screen "08 BTCS MAIN" 1280x800, template "Template"
   Rectangle "Rectangle_2" at 150,205 size 480x40
      Appearance <- "2102_TIME_CALCS_DB_DE_OX_TMR_DN"
   TextField "Text field_7" at 155,210 size 200x30; Text 'De-Oxygenate Time :'
   IOField "I/O field_3" at 360,210 size 60x30; FormatPattern 999
      ProcessValue <- "2110_BTCS_CNTRL_DB_DE_OX_HRS"
   TextField "Text field_8" at 420,210 size 60x30; Text 'Hours'
   IOField "I/O field_4" at 485,210 size 60x30; FormatPattern 99
      ProcessValue <- "2110_BTCS_CNTRL_DB_DE_OX_MINS"
   TextField "Text field_9" at 545,210 size 80x30; Text 'Minutes'
   Rectangle "Rectangle_3" at 150,250 size 480x40
      Appearance <- "2102_TIME_CALCS_DB_DWELL_TMR_DN"
   TextField "Text field_10" at 155,255 size 200x30; Text 'Dwell Time :'
   IOField "I/O field_5" at 360,255 size 60x30; FormatPattern 999
      ProcessValue <- "2110_BTCS_CNTRL_DB_DWELL_HRS"
   TextField "Text field_11" at 420,255 size 60x30; Text 'Hours'
   IOField "I/O field_6" at 485,255 size 60x30; FormatPattern 99
      ProcessValue <- "2110_BTCS_CNTRL_DB_DWELL_MINS"
   TextField "Text field_12" at 545,255 size 80x30; Text 'Minutes'
   Rectangle "Rectangle_4" at 150,295 size 480x40
      Appearance <- "2102_TIME_CALCS_DB_RE_OX_TMR_DN"
   TextField "Text field_13" at 155,300 size 200x30; Text 'Re-Oxygenate Time :'
   IOField "I/O field_7" at 360,300 size 60x30; FormatPattern 999
      ProcessValue <- "2110_BTCS_CNTRL_DB_RE_OX_HRS"
   TextField "Text field_14" at 420,300 size 60x30; Text 'Hours'
   IOField "I/O field_8" at 485,300 size 60x30; FormatPattern 99
      ProcessValue <- "2110_BTCS_CNTRL_DB_RE_OX_MINS"
   TextField "Text field_15" at 545,300 size 80x30; Text 'Minutes'
   Rectangle "Rectangle_5" at 150,340 size 480x40
      Appearance <- "2102_TIME_CALCS_DB_POST_DWELL_TMR_DN"
   TextField "Text field_16" at 155,345 size 200x30; Text 'Post-Dwell Time :'
   IOField "I/O field_9" at 360,345 size 60x30; FormatPattern 999
      ProcessValue <- "2110_BTCS_CNTRL_DB_POST_DWELL_HRS"
   TextField "Text field_17" at 420,345 size 60x30; Text 'Hours'
   IOField "I/O field_10" at 485,345 size 60x30; FormatPattern 99
      ProcessValue <- "2110_BTCS_CNTRL_DB_POST_DWELL_MINS"
   TextField "Text field_18" at 545,345 size 80x30; Text 'Minutes'
   Rectangle "Rectangle_6" at 640,205 size 480x40
      Appearance <- "2102_TIME_CALCS_DB_DE_OX_SP_TMR_DN"
   TextField "Text field_19" at 645,210 size 200x30; Text 'At De-Ox Setpoint :'
   IOField "I/O field_11" at 850,210 size 60x30; FormatPattern 999
      ProcessValue <- "2110_BTCS_CNTRL_DB_DE_OX_SP_HRS"
   TextField "Text field_20" at 910,210 size 60x30; Text 'Hours'
   IOField "I/O field_12" at 975,210 size 60x30; FormatPattern 99
      ProcessValue <- "2110_BTCS_CNTRL_DB_DE_OX_SP_MINS"
   TextField "Text field_21" at 1035,210 size 80x30; Text 'Minutes'
   Rectangle "Rectangle_7" at 640,295 size 480x40
      Appearance <- "2102_TIME_CALCS_DB_RE_OX_SP_TMR_DN"
   TextField "Text field_22" at 645,300 size 200x30; Text 'At Re-Ox Setpoint :'
   IOField "I/O field_13" at 850,300 size 60x30; FormatPattern 999
      ProcessValue <- "2110_BTCS_CNTRL_DB_RE_OX_SP_HRS"
   TextField "Text field_23" at 910,300 size 60x30; Text 'Hours'
   IOField "I/O field_14" at 975,300 size 60x30; FormatPattern 99
      ProcessValue <- "2110_BTCS_CNTRL_DB_RE_OX_SP_MINS"
   TextField "Text field_24" at 1035,300 size 80x30; Text 'Minutes'
   TextField "Text field_25" at 155,435 size 200x30; Text 'Total Sequence Time:'
   IOField "I/O field_15" at 360,435 size 60x30; FormatPattern 999
      ProcessValue <- "2110_BTCS_CNTRL_DB_TOT_SEQ_HRS"
   TextField "Text field_26" at 420,435 size 60x30; Text 'Hours'
   IOField "I/O field_16" at 485,435 size 60x30; FormatPattern 99
      ProcessValue <- "2110_BTCS_CNTRL_DB_TOT_SEQ_MINS"
   TextField "Text field_27" at 545,435 size 80x30; Text 'Minutes'
   TextField "Text field_28" at 155,625 size 200x30; Text 'Remaining Time:'
   IOField "I/O field_17" at 360,625 size 60x30; FormatPattern 999
      ProcessValue <- "2110_BTCS_CNTRL_DB_RMNG_SEQ_HRS"
   TextField "Text field_29" at 420,625 size 60x30; Text 'Hours'
   IOField "I/O field_18" at 485,625 size 60x30; FormatPattern 99
      ProcessValue <- "2110_BTCS_CNTRL_DB_RMNG_SEQ_MINS"
   TextField "Text field_30" at 545,625 size 80x30; Text 'Minutes'
   TextField "Text field_61" at 150,575 size 480x35; Text 'INPUT SALINITY'
      Visibility <- "2068_Sys_Status_Data_SAL_VALID"
   TextField "Text field_60" at 150,575 size 480x35; Text 'SALINITY ACCEPTED'
      Visibility <- "2068_Sys_Status_Data_SAL_VALID"
   Button "HmiScreenItemData_1" at 10,10 size 160x50; TextOn 'Back'; TextOff 'Main Index'
      on Release: ActivateScreen("02 Main Index", 0)
   TextField "Text field_1" at 324,55 size 640x35; Text 'BASIC BARGE TWO TANK CONTROL SYSTEM'
   Button "HmiScreenItemData_2" at 1127,4 size 149x50; TextOn 'Back'; TextOff 'Enable'
      on Press: ResetBit("80_From_HMI_RUN_BWTS"); SetBit("80_From_HMI_RUN_BTCS")
      Visibility <- "80_From_HMI_RUN_BTCS"
   Button "HmiScreenItemData_3" at 1127,56 size 149x50; TextOn 'Back'; TextOff 'Disable'
      on Press: ResetBit("80_From_HMI_RUN_BTCS"); SetBit("80_From_HMI_RUN_BWTS")
      Visibility <- "80_From_HMI_RUN_BTCS"
   TextField "Text field_2" at 484,85 size 320x35; Text 'BTCS ENABLED'
      Visibility <- "80_From_HMI_RUN_BTCS"
   TextField "Text field_3" at 484,85 size 320x35; Text 'BTCS DISABLED'
      Visibility <- "80_From_HMI_RUN_BTCS"
   Button "Button_2" at 10,70 size 160x50; TextOn 'User Account'; TextOff 'Alarm Log'; Authorization "User administration"
      on Release: ActivateScreen("04 Alarm Log", 0)
   Group "Group_1" at 150,205 size 480x40
   Group "Group_2" at 150,250 size 480x40
   Group "Group_3" at 150,295 size 480x40
   Group "Group_4" at 150,340 size 480x40
   Group "Group_5" at 640,205 size 480x40
   Group "Group_6" at 640,295 size 480x40
   Group "Group_7" at 150,430 size 480x40
   Group "Group_8" at 150,620 size 480x40
   TextField "Text field_31" at 1005,150 size 120x30; Text 'SETUP'
   TextField "Text field_32" at 1005,420 size 120x30; Text 'CONTROL'
   Button "Button_1" at 150,520 size 230x50; TextOff 'ACCEPT & LAUNCH'
      on Release: ResetBit("2110_BTCS_CNTRL_DB_START_SEQ")
      on Press: SetBit("2110_BTCS_CNTRL_DB_START_SEQ")
      Appearance <- "2110_BTCS_CNTRL_DB_BTCS_STATE"
      Visibility <- "2102_TIME_CALCS_DB_TIMES_VALID"
   SymbolicIOField "Symbolic I/O field_1" at 640,480 size 480x30; TextOn '1'; TextOff '0'; TextList "STATE LIST BTCS"
      ProcessValue <- "2110_BTCS_CNTRL_DB_BTCS_STATE"
   TextField "Text field_33" at 150,480 size 480x35; Text 'TIMES NOT VALID'
      Visibility <- "2102_TIME_CALCS_DB_TIMES_VALID"
   TextField "Text field_34" at 150,480 size 480x35; Text 'TIMES VALID'
      Visibility <- "2102_TIME_CALCS_DB_TIMES_VALID"
   SymbolicIOField "Symbolic I/O field_2" at 640,580 size 480x30; TextOn '1'; TextOff '0'; TextList "STEP LIST BTCS"
      ProcessValue <- "2110_BTCS_CNTRL_DB_BTCS_STEP"
   Button "HmiScreenItemData_4" at 1127,108 size 149x50; TextOn 'Back'; TextOff 'Master Reset'
      on Press: ResetBit("2110_BTCS_CNTRL_DB_RESET_ALL"); SetBit("2110_BTCS_CNTRL_DB_RESET_ALL")
      Visibility <- "80_From_HMI_RUN_BTCS"
   SymbolicIOField "Symbolic I/O field_3" at 360,700 size 140x30; TextOn '1'; TextOff '0'; TextList "Port Tank"
      ProcessValue <- "2110_BTCS_CNTRL_DB_PORT_TANK_STS"
   Button "Button_4" at 150,700 size 180x30; TextOff 'Port Tank'
      on Press: InvertBit("2110_BTCS_CNTRL_DB_PORT_TANK_STS")
      Appearance <- "2110_BTCS_CNTRL_DB_PORT_TANK_STS"
   TextField "Text field_35" at 1025,690 size 100x30; Text 'TANKS'
   SymbolicIOField "Symbolic I/O field_4" at 360,740 size 140x30; TextOn '1'; TextOff '0'; TextList "Port Tank"
      ProcessValue <- "2110_BTCS_CNTRL_DB_STBD_TANK_STS"
   Button "Button_5" at 150,740 size 180x30; TextOff 'Starboard Tank'
      on Press: InvertBit("2110_BTCS_CNTRL_DB_STBD_TANK_STS")
      Appearance <- "2110_BTCS_CNTRL_DB_STBD_TANK_STS"
   TextField "Text field_37" at 515,700 size 60x30; Text 'O2 :'
   IOField "I/O field_20" at 575,700 size 60x30; FormatPattern 99.99
      ProcessValue <- "20_TANKS_IP_DATA_RIO_02_FIRST_TANK_BWT_DO"
   TextField "Text field_36" at 640,700 size 60x30; Text 'ph :'
   IOField "I/O field_19" at 700,700 size 60x30; FormatPattern 99.99
      ProcessValue <- "20_TANKS_IP_DATA_RIO_02_FIRST_TANK_BWT_PH"
   TextField "Text field_38" at 775,700 size 65x30; Text 'Temp :'
   IOField "I/O field_21" at 840,700 size 60x30; FormatPattern 99.99
      ProcessValue <- "20_TANKS_IP_DATA_RIO_02_FIRST_TANK_BWT_TEMP"
   TextField "Text field_39" at 910,700 size 65x30; Text 'Level :'
   IOField "I/O field_22" at 975,700 size 60x30; FormatPattern 99.9
      ProcessValue <- "20_TANKS_IP_DATA_RIO_02_FIRST_TANK_BWT_LEVEL"
   TextField "Text field_40" at 515,740 size 60x30; Text 'O2 :'
   IOField "I/O field_23" at 575,740 size 60x30; FormatPattern 99.99
      ProcessValue <- "20_TANKS_IP_DATA_RIO_02_SECOND_TANK_BWT_DO"
   TextField "Text field_41" at 640,740 size 60x30; Text 'ph :'
   IOField "I/O field_24" at 700,740 size 60x30; FormatPattern 99.99
      ProcessValue <- "20_TANKS_IP_DATA_RIO_02_SECOND_TANK_BWT_PH"
   TextField "Text field_42" at 775,740 size 65x30; Text 'Temp :'
   IOField "I/O field_25" at 840,740 size 60x30; FormatPattern 99.99
      ProcessValue <- "20_TANKS_IP_DATA_RIO_02_SECOND_TANK_BWT_TEMP"
   TextField "Text field_43" at 910,740 size 65x30; Text 'Level :'
   IOField "I/O field_26" at 975,740 size 60x30; FormatPattern 99.9
      ProcessValue <- "20_TANKS_IP_DATA_RIO_02_SECOND_TANK_BWT_LEVEL"
   Group "Group" at 150,160 size 480x40
   Group "Group_9" at 150,160 size 480x40
   Group "Group_10" at 150,340 size 480x40
   Group "Group_12" at 150,295 size 480x40
   Group "Group_13" at 640,205 size 480x40
   Group "Group_14" at 150,250 size 480x40
   Group "Group_15" at 150,205 size 480x40
   Group "Group_16" at 640,295 size 480x40
   Rectangle "Rectangle_15" at 249,485 size 303x130
      Visibility <- "2100_AUTO_SEQ_DB_SEQ_RNG"
   Button "Button_3" at 400,520 size 230x50; TextOff 'ABORT - STOP'
      on Release: ResetBit("2110_BTCS_CNTRL_DB_STOP_SEQ")
      on Press: SetBit("2110_BTCS_CNTRL_DB_STOP_SEQ")
      Appearance <- "2110_BTCS_CNTRL_DB_BTCS_STATE"
   Group "Group_17" at 640,250 size 480x40
   Group "Group_18" at 640,250 size 480x40
   Group "Group_11" at 647,276 size 480x40
   Group "Group_19" at 1083,420 size 47x365
   Rectangle "Rectangle_1" at 150,160 size 480x40
      Appearance <- "2102_TIME_CALCS_DB_PRE_DWELL_TMR_DN"
   TextField "Text field_4" at 155,165 size 200x30; Text 'Pre-Dwell Time :'
   IOField "I/O field_1" at 360,165 size 60x30; FormatPattern 999
      ProcessValue <- "2110_BTCS_CNTRL_DB_PRE_DWELL_HRS"
   TextField "Text field_5" at 420,165 size 60x30; Text 'Hours'
   IOField "I/O field_2" at 485,165 size 60x30; FormatPattern 99
      ProcessValue <- "2110_BTCS_CNTRL_DB_PRE_DWELL_MINS"
   TextField "Text field_6" at 545,165 size 80x30; Text 'Minutes'
   Rectangle "Rectangle_13" at 150,160 size 480x40
      Visibility <- "2100_AUTO_SEQ_DB_SEQ_RNG"
      Appearance <- "2102_TIME_CALCS_DB_PRE_DWELL_TMR_DN"
   TextField "Text field_44" at 155,165 size 310x30; Text 'Pre-Dwell Time Remaining :'
      Visibility <- "2100_AUTO_SEQ_DB_SEQ_RNG"
   IOField "I/O field_28" at 465,165 size 80x30; FormatPattern 999999
      Visibility <- "2100_AUTO_SEQ_DB_SEQ_RNG"
      ProcessValue <- "2102_TIME_CALCS_DB_PRE_DWELL_MINS_RMNG"
   TextField "Text field_46" at 545,165 size 80x30; Text 'Minutes'
      Visibility <- "2100_AUTO_SEQ_DB_SEQ_RNG"
   Rectangle "Rectangle_14" at 150,340 size 480x40
      Visibility <- "2100_AUTO_SEQ_DB_SEQ_RNG"
      Appearance <- "2102_TIME_CALCS_DB_POST_DWELL_TMR_DN"
   TextField "Text field_45" at 155,345 size 310x30; Text 'Post-Dwell Time Remaining :'
      Visibility <- "2100_AUTO_SEQ_DB_SEQ_RNG"
   IOField "I/O field_27" at 465,345 size 80x30; FormatPattern 999999
      ProcessValue <- "2102_TIME_CALCS_DB_POST_DWELL_MINS_RMNG"
      Visibility <- "2100_AUTO_SEQ_DB_SEQ_RNG"
   TextField "Text field_47" at 545,345 size 80x30; Text 'Minutes'
      Visibility <- "2100_AUTO_SEQ_DB_SEQ_RNG"
   Rectangle "Rectangle_16" at 150,295 size 480x40
      Visibility <- "2100_AUTO_SEQ_DB_SEQ_RNG"
      Appearance <- "2102_TIME_CALCS_DB_RE_OX_TMR_DN"
   TextField "Text field_50" at 155,300 size 310x30; Text 'Re-Oxygenate Time Remaining :'
      Visibility <- "2100_AUTO_SEQ_DB_SEQ_RNG"
   IOField "I/O field_30" at 465,300 size 80x30; FormatPattern 999999
      ProcessValue <- "2102_TIME_CALCS_DB_RE_OX_MINS_RMNG"
      Visibility <- "2100_AUTO_SEQ_DB_SEQ_RNG"
   TextField "Text field_51" at 545,300 size 80x30; Text 'Minutes'
      Visibility <- "2100_AUTO_SEQ_DB_SEQ_RNG"
   Rectangle "Rectangle_17" at 640,205 size 480x40
      Visibility <- "2100_AUTO_SEQ_DB_SEQ_RNG"
      Appearance <- "2102_TIME_CALCS_DB_DE_OX_SP_TMR_DN"
   TextField "Text field_52" at 645,210 size 310x30; Text 'At De-Ox Time Remaining :'
      Visibility <- "2100_AUTO_SEQ_DB_SEQ_RNG"
   IOField "I/O field_31" at 955,210 size 80x30; FormatPattern 999999
      ProcessValue <- "2102_TIME_CALCS_DB_DE_OX_SP_MINS_RMNG"
      Visibility <- "2100_AUTO_SEQ_DB_SEQ_RNG"
   TextField "Text field_53" at 1035,210 size 80x30; Text 'Minutes'
      Visibility <- "2100_AUTO_SEQ_DB_SEQ_RNG"
   Rectangle "Rectangle_18" at 150,250 size 480x40
      Visibility <- "2100_AUTO_SEQ_DB_SEQ_RNG"
      Appearance <- "2102_TIME_CALCS_DB_DWELL_TMR_DN"
   TextField "Text field_54" at 155,255 size 310x30; Text 'Dwell Time Remaining :'
      Visibility <- "2100_AUTO_SEQ_DB_SEQ_RNG"
   IOField "I/O field_32" at 465,255 size 80x30; FormatPattern 999999
      ProcessValue <- "2102_TIME_CALCS_DB_DWELL_MINS_RMNG"
      Visibility <- "2100_AUTO_SEQ_DB_SEQ_RNG"
   TextField "Text field_55" at 545,255 size 80x30; Text 'Minutes'
      Visibility <- "2100_AUTO_SEQ_DB_SEQ_RNG"
   Rectangle "Rectangle_19" at 150,205 size 480x40
      Visibility <- "2100_AUTO_SEQ_DB_SEQ_RNG"
      Appearance <- "2102_TIME_CALCS_DB_DE_OX_TMR_DN"
   TextField "Text field_56" at 155,210 size 310x30; Text 'De-Oxygenate Time Remaining :'
      Visibility <- "2100_AUTO_SEQ_DB_SEQ_RNG"
   IOField "I/O field_33" at 465,210 size 80x30; FormatPattern 999999
      ProcessValue <- "2102_TIME_CALCS_DB_DE_OX_MINS_RMNG"
      Visibility <- "2100_AUTO_SEQ_DB_SEQ_RNG"
   TextField "Text field_57" at 545,210 size 80x30; Text 'Minutes'
      Visibility <- "2100_AUTO_SEQ_DB_SEQ_RNG"
   Rectangle "Rectangle_20" at 640,295 size 480x40
      Visibility <- "2100_AUTO_SEQ_DB_SEQ_RNG"
      Appearance <- "2102_TIME_CALCS_DB_RE_OX_SP_TMR_DN"
   TextField "Text field_58" at 645,300 size 310x30; Text 'At Re-Ox Time Remaining :'
      Visibility <- "2100_AUTO_SEQ_DB_SEQ_RNG"
   IOField "I/O field_34" at 955,300 size 80x30; FormatPattern 999999
      ProcessValue <- "2102_TIME_CALCS_DB_RE_OX_SP_MINS_RMNG"
      Visibility <- "2100_AUTO_SEQ_DB_SEQ_RNG"
   TextField "Text field_59" at 1035,300 size 80x30; Text 'Minutes'
      Visibility <- "2100_AUTO_SEQ_DB_SEQ_RNG"
   Rectangle "Rectangle_22" at 647,276 size 480x40
      Visibility <- "2100_AUTO_SEQ_DB_SEQ_RNG"
      Appearance <- "2102_TIME_CALCS_DB_RE_OX_SP_TMR_DN"
   TextField "Text field_49" at 652,281 size 310x30; Text 'Salinity Value :'
      Visibility <- "2100_AUTO_SEQ_DB_SEQ_RNG"
   IOField "I/O field_36" at 962,281 size 90x30; FormatPattern 99.9; Unit psu
      Visibility <- "2100_AUTO_SEQ_DB_SEQ_RNG"
      ProcessValue <- "80_From_HMI_SAL_VALUE"
   Rectangle "Rectangle_21" at 640,250 size 480x40
      Appearance <- "2068_Sys_Status_Data_SAL_VALID"
   TextField "Text field_48" at 645,255 size 200x30; Text 'Set Salinity Value :'
   IOField "I/O field_29" at 850,255 size 90x30; FormatPattern 99.9; Unit psu
      ProcessValue <- "80_From_HMI_SAL_VALUE"
   Button "HmiScreenItemData_5" at 955,255 size 150x30; TextOn 'Back'; TextOff 'Confirm Salinity'
      on Press: function_b14e0dd5("80_From_HMI_SAL_CNFRM", 0)
   Rectangle "Rectangle_23" at 640,250 size 480x40
      Visibility <- "2068_Sys_Status_Data_SAL_CNF_CHK"
   TextField "Text field_62" at 645,255 size 250x30; Text 'Salinity Value < 1 Confirm? :'
      Visibility <- "2068_Sys_Status_Data_SAL_CNF_CHK"
   Button "Button_6" at 910,255 size 80x30; TextOff 'YES'
      on Press: function_b14e0dd5("80_From_HMI_LOW_SAL_ACPT", 0)
      Visibility <- "2068_Sys_Status_Data_SAL_CNF_CHK"
   Button "Button_7" at 1020,255 size 80x30; TextOff 'NO'
      on Press: function_b14e0dd5("80_From_HMI_LOW_SAL_RJCT", 0)
      Visibility <- "2068_Sys_Status_Data_SAL_CNF_CHK"
   Rectangle "Rectangle_24" at 1083,420 size 47x365
      Visibility <- "2068_Sys_Status_Data_SAL_CNF_CHK"
   TextField "Text field_65" at 1084,450 size 46x80; Text '!!! WARNING Salinity < 1 Outside Of Certified Range !!!'
      Visibility <- "2068_Sys_Status_Data_SAL_CNF_CHK"
   TextField "Text field_66" at 1084,550 size 46x80; Text 'Confirming Above Means :'
      Visibility <- "2068_Sys_Status_Data_SAL_CNF_CHK"
   TextField "Text field_67" at 1084,650 size 46x80; Text '!!! User Takes Responsability For This Action !!!'
      Visibility <- "2068_Sys_Status_Data_SAL_CNF_CHK"

screen "09 Sys Config" 1280x800, template "Template"
   Circle "Circle_2" at 221,236 size 29x29
      Appearance <- "82_To_HMI_CRNT_MODE_IGG"
   Button "HmiScreenItemData_1" at 1,1 size 150x43; TextOn 'Back'; TextOff 'Main Index'
      on Release: ActivateScreen("02 Main Index", 0)
   Button "HmiScreenItemData_8" at 44,70 size 230x29; TextOn 'Back'; TextOff 'IGG Mode of Operation'
   Circle "Circle_1" at 221,177 size 29x29
      Appearance <- "82_To_HMI_CRNT_MODE_IGG"
   Button "HmiScreenItemData_4" at 50,167 size 150x51; TextOn 'Back'; TextOff 'Manual'; Authorization "Operating Mode"
      on Press: function_b14e0dd5("80_From_HMI_Request_Manual(1)", 0)
   Circle "Circle_9" at 221,116 size 29x29
      Appearance <- "82_To_HMI_CRNT_MODE_IGG"
   TextField "Text field_13" at 293,112 size 93x21; Text 'Description'
   IOField "I/O field_13" at 463,189 size 226x30; FormatPattern 9999999999999999999999999999999999999999
      ProcessValue <- "db_time_sync_time_system_READ"
   Button "HmiScreenItemData_26" at 284,70 size 421x29; TextOn 'Back'; TextOff 'Time Setting'
   Button "HmiScreenItemData_24" at 291,231 size 166x30; TextOn 'Back'; TextOff 'Set System Time'; Authorization "Parameter Change"
      on Activate: function_cbf290fd(0, 0)
   Button "HmiScreenItemData_16" at 894,69 size 187x29; TextOn 'Back'; TextOff 'IO'
   Button "HmiScreenItemData_2" at 719,69 size 163x29; TextOn 'Back'; TextOff 'Runtime'
   Button "HmiScreenItemData_10" at 725,107 size 150x51; TextOn 'Back'; TextOff 'Reset AUTO'; Authorization "User administration"
      on Press: function_b14e0dd5("80_From_HMI_RST_AUT_SEQ(1)", 0)
      Appearance <- "80_From_HMI_RST_AUT_SEQ(1)"
   DateTimeField "Date/time field_1" at 463,231 size 226x30; Authorization "Parameter Change"
   TextField "Text field_14" at 314,195 size 142x20; Text 'System Time (UTC)'
   Button "HmiScreenItemData_23" at 50,106 size 150x51; TextOn 'Back'; TextOff 'Full Automation'; Authorization "Operating Mode"
      on Press: function_b14e0dd5("80_From_HMI_Request_Auto(1)", 0)
   Button "HmiScreenItemData_3" at 1129,1 size 150x43; TextOn 'I&A Compressor Ok'; TextOff 'Back'
      on Release: function_efd93a16()
   Button "HmiScreenItemData_7" at 50,228 size 150x51; TextOn 'Back'; TextOff 'FAT Mode'; Authorization "User administration"
      on Press: InvertBit("80_From_HMI_FAT_Mode"); function_b14e0dd5("80_From_HMI_Request_Auto(1)", 0)
   Button "HmiScreenItemData_11" at 725,232 size 150x51; TextOn 'Back'; TextOff 'IGG Standalone'; Authorization "Operating Mode"
      on Press: InvertBit("80_From_HMI_IGG_STND_ALN")
      Appearance <- "80_From_HMI_IGG_STND_ALN"
   Button "HmiScreenItemData_12" at 910,100 size 150x51; TextOn 'Back'; TextOff 'P301 Present'; Authorization "Operating Mode"; TextList "P301 Present"
      on Press: InvertBit("80_From_HMI_P301_PRSNT(1)")
      Appearance <- "80_From_HMI_P301_PRSNT(1)"
      ProcessValue <- "80_From_HMI_P301_PRSNT(1)"
   Button "HmiScreenItemData_13" at 910,155 size 150x51; TextOn 'Back'; TextOff 'CV312 Present'; Authorization "User administration"; TextList "CV312 Present"
      on Press: InvertBit("80_From_HMI_CV312_PRSNT")
      Appearance <- "80_From_HMI_CV312_PRSNT"
      ProcessValue <- "80_From_HMI_CV312_PRSNT"
   Button "HmiScreenItemData_14" at 910,212 size 150x51; TextOn 'Back'; TextOff 'CV431 Present'; Authorization "Operating Mode"; TextList "CV431 Present"
      on Press: InvertBit("80_From_HMI_CV431_PRSNT")
      Appearance <- "80_From_HMI_CV431_PRSNT"
      ProcessValue <- "80_From_HMI_CV431_PRSNT"
   Button "HmiScreenItemData_15" at 910,269 size 150x51; TextOn 'Back'; TextOff 'CV432 Present'; Authorization "Operating Mode"; TextList "CV432 Present"
      on Press: InvertBit("80_From_HMI_CV432_PRSNT")
      Appearance <- "80_From_HMI_CV432_PRSNT"
      ProcessValue <- "80_From_HMI_CV432_PRSNT"
   Button "HmiScreenItemData_18" at 725,166 size 150x51; TextOn 'Back'; TextOff 'Silence Buzzer'; Authorization "User administration"
      on Press: function_b14e0dd5("80_From_HMI_SLNCE_BZR", 0)
      Appearance <- "80_From_HMI_SLNCE_BZR"
   AlarmView "Alarm view_1" at 0,777 size 1280x23
   IOField "I/O field_9" at 1024,352 size 60x30; Authorization "Commissioning"; FormatPattern 99; Unit  s
      ProcessValue <- "80_From_HMI_Beacon frequency"
   IOField "I/O field_10" at 1025,389 size 60x30; Authorization "Commissioning"; FormatPattern 99; Unit  min
      ProcessValue <- "80_From_HMI_Buzzer reset time"
   TextField "Text field_9" at 895,358 size 138x20; Text 'Beacon frequency'
   TextField "Text field_10" at 895,394 size 100x20; Text 'Buzzer reset'

screen "Main Page" 1280x800, template "Template"
   GraphicView "Graphic view_49" at 158,415 size 30x45; Picture "Graphic_72"
   GraphicView "Graphic view_20" at 140,368 size 380x356; Picture "IGG_6"
   GraphicView "Graphic view_62" at 134,449 size 92x8; Picture "Graphic_20"
   GraphicView "Graphic view_5" at 464,423 size 90x19; Picture "Graphic_82"
   GraphicView "Graphic view_41" at 228,459 size 9x40; Picture "Graphic_57"
   GraphicView "Graphic view_40" at 222,449 size 15x13; Picture "Graphic_41"
   GraphicView "Graphic view_21" at 210,503 size 17x7; Picture "Graphic_63"
   GraphicView "Graphic view_22" at 207,499 size 8x9; Picture "Graphic_64"
   GraphicView "Graphic view_23" at 206,399 size 6x104; Picture "Graphic_70"
   GraphicView "Graphic view_39" at 138,535 size 6x7; Picture "Graphic_70"
   GraphicView "Graphic view_38" at 139,539 size 7x9; Picture "Graphic_64"
   GraphicView "Graphic view_18" at 204,397 size 9x10; Picture "Graphic_67"
   Group "Group_3" at 158,415 size 30x41; Picture "Graphic_72"
   GraphicView "Graphic view_65" at 144,542 size 8x6; Picture "Graphic_63"
   GraphicView "Graphic view_69" at 295,453 size 14x15; Picture "Graphic_36"
   GraphicView "Graphic view_70" at 335,462 size 14x15; Picture "Graphic_36"
   GraphicView "Graphic view_71" at 251,443 size 14x17; Picture "Graphic_79"
   GraphicView "Graphic view_36" at 517,373 size 35x50; Picture "Graphic_108"
   GraphicView "Graphic view_4" at 333,376 size 31x49; Picture "Graphic_108"
   GraphicView "Graphic view_72" at 387,407 size 14x17; Picture "Graphic_36"
   GraphicView "Graphic view_37" at 136,525 size 8x11; Picture "Graphic_67"
   GraphicView "Graphic view_89" at 440,407 size 14x17; Picture "Graphic_36"
   Line "Line_4" at 226,517 size 2x15
      Visibility <- "14_DQ_Data_X001ControlOut"
   GraphicView "Graphic view_84" at 215,511 size 27x55; Picture "Graphic_129"
      Visibility <- "102_Pilot_Burner_DB_FLM_DET"
   GraphicView "Graphic view_90" at 488,409 size 14x15; Picture "Graphic_36"
   GraphicView "Graphic view_1" at 342,415 size 18x41; Picture "Graphic_17"
   GraphicView "Graphic view_60" at 526,412 size 18x41; Picture "Graphic_17"
   GraphicView "Graphic view_82" at 210,499 size 167x147; Picture "Graphic_130"
      Visibility <- "103_Main_Burner_DB_DN_OK(1)"
   IOField "I/O field_17" at 231,558 size 46x17; FormatPattern 999; Unit %
      ProcessValue <- "12_AI_Data_FD001FlameSignalIn"
      Visibility <- "10 DI_DATA_FD001_OK"
   GraphicView "Graphic view_63" at 133,396 size 75x7; Picture "Graphic_63"
   Group "Group_10" at 659,340 size 26x47; Picture "Graphic_148"
   Group "Group_11" at 649,372 size 56x37; Picture "Graphic_224"
   GraphicView "Graphic view_25" at 659,340 size 25x46; Picture "Graphic_148"
   GraphicView "Graphic view_26" at 649,373 size 55x36; Picture "Graphic_224"
   GraphicView "Graphic view_27" at 569,502 size 205x15; Picture "Graphic_232"
   GraphicView "Graphic view_3" at 78,471 size 64x14; Picture "Graphic_82"
   GraphicView "Graphic view_19" at 776,616 size 64x10; Picture "Graphic_82"
   GraphicIOField "Graphic I/O field_2" at 0,485 size 128x131; PictureList "IA Compressor_1"
      ProcessValue <- "82_To_HMI_CA Blower Animation"
   GraphicView "Graphic view_7" at 700,602 size 119x212; Picture "Graphic_150"
   Group "Group" at 133,368 size 421x356; Picture "Graphic_20"
   GraphicView "Graphic view_2" at 821,493 size 449x266; Picture "Graphic_185"
   GraphicView "Graphic view_6" at 68,470 size 18x21; Picture "Graphic_66"
   GraphicView "Graphic view_8" at 41,328 size 96x93; Picture "Graphic_246"
   GraphicView "Graphic view_14" at 630,544 size 17x40; Picture "Graphic_271"
   GraphicView "Graphic view_15" at 570,390 size 205x15; Picture "Graphic_232"
   GraphicView "Graphic view_16" at 561,391 size 26x27; Picture "Graphic_178"
   GraphicView "Graphic view_17" at 757,380 size 17x35; Picture "Graphic_280"
   GraphicView "Graphic view_9" at 525,539 size 156x153; Picture "Graphic_251"
   GraphicView "Graphic view_24" at 561,407 size 14x167; Picture "Graphic_231"
   GraphicView "Graphic view_11" at 555,635 size 21x22; Picture "Graphic_265"
   GraphicView "Graphic view_12" at 555,653 size 29x31; Picture "Graphic_266"
   GraphicView "Graphic view_13" at 572,667 size 133x18; Picture "Graphic_232"
   GraphicView "Graphic view_10" at 549,422 size 26x38; Picture "Graphic_169"
   Group "Group_12" at 649,340 size 56x69; Picture "Graphic_148"
   GraphicView "Graphic view_28" at 756,492 size 17x35; Picture "Graphic_280"
   Group "Group_4" at 648,452 size 56x69; Picture "Graphic_148"
   Group "Group_1" at 658,452 size 26x47; Picture "Graphic_148"
   Group "Group_2" at 648,484 size 56x37; Picture "Graphic_224"
   GraphicView "Graphic view_29" at 658,452 size 25x46; Picture "Graphic_148"
   GraphicView "Graphic view_30" at 648,485 size 55x36; Picture "Graphic_224"

screen "IGG Analogue Inputs" 1280x800, template "Template"
   on GenerateScreen: "TitleUpdater"()
   Button "HmiScreenItemData_1" at 1,1 size 150x43; TextOn 'Back'; TextOff 'Commissioning'
      on Release: ActivateScreen("Commissioning Main Page", 0)
   TextField "Text field_82" at 60,150 size 220x22; Text 'PIT-102 - CA Pressure (Pre-Ignition)'
   TextField "Text field_90" at 286,124 size 64x20; Text 'Reading'
   IOField "I/O field_2" at 287,150 size 70x22; FormatPattern 9999; Unit  mBar
      ProcessValue <- "12_AI_Data_PIT102_SCALED(1)"
   TextField "Text field_1" at 359,124 size 68x20; Text 'Low Low'
   IOField "I/O field_1" at 361,150 size 60x22; Authorization "Parameter Change"; FormatPattern 9999
      ProcessValue <- "84_Setpoints_PIT102_Pilot_LowLow"
   TextField "Text field_2" at 442,124 size 37x20; Text 'Low'
   IOField "I/O field_3" at 429,150 size 60x22; Authorization "Parameter Change"; FormatPattern 9999
      ProcessValue <- "84_Setpoints_PIT102_Pilot_Low"
   TextField "Text field_3" at 509,124 size 37x20; Text 'High'
   IOField "I/O field_4" at 497,150 size 60x22; Authorization "Parameter Change"; FormatPattern 9999
      ProcessValue <- "84_Setpoints_PIT102_Pilot_High"
   TextField "Text field_4" at 561,124 size 74x20; Text 'High High'
   IOField "I/O field_5" at 565,150 size 60x22; Authorization "Parameter Change"; FormatPattern 9999
      ProcessValue <- "84_Setpoints_PIT102_Pilot_HighHigh"
   TextField "Text field_5" at 434,100 size 76x20; Text 'Setpoints'
   TextField "Text field_6" at 7,150 size 53x22; Text 'IW112'
   TextField "Text field_7" at 60,270 size 220x22; Text 'TIT-401 - IG Temperature'
   IOField "I/O field_6" at 287,270 size 70x22; FormatPattern s999.9; Unit  °C
      ProcessValue <- "12_AI_Data_TIT401_SCALED"
   IOField "I/O field_7" at 361,270 size 60x22; FormatPattern s999.9
   IOField "I/O field_8" at 429,270 size 60x22; FormatPattern s999.9
   IOField "I/O field_9" at 497,270 size 60x22; Authorization "Parameter Change"; FormatPattern s999.9
      ProcessValue <- "84_Setpoints_TIT401_High"
   IOField "I/O field_10" at 565,270 size 60x22; Authorization "Parameter Change"; FormatPattern s999.9
      ProcessValue <- "84_Setpoints_TIT401_HighHigh"
   TextField "Text field_8" at 7,270 size 53x22; Text 'IW114'
   TextField "Text field_9" at 60,310 size 220x22; Text 'PIT-402 - IG Outlet Pres. (Pre-Ignitn.)'
   IOField "I/O field_11" at 287,310 size 70x22; FormatPattern 9999; Unit  mBar
      ProcessValue <- "12_AI_Data_PIT402_SCALED"
   IOField "I/O field_12" at 361,310 size 60x22; Authorization "Parameter Change"; FormatPattern 9999
      ProcessValue <- "84_Setpoints_PIT402_Pilot_LowLow"
   IOField "I/O field_13" at 429,310 size 60x22; Authorization "Parameter Change"; FormatPattern 9999
      ProcessValue <- "84_Setpoints_PIT402_Pilot_Low"
   IOField "I/O field_14" at 497,310 size 60x22; Authorization "Parameter Change"; FormatPattern 9999
      ProcessValue <- "84_Setpoints_PIT402_Pilot_High"
   IOField "I/O field_15" at 565,310 size 60x22; Authorization "Parameter Change"; FormatPattern 9999
      ProcessValue <- "84_Setpoints_PIT402_Pilot_HighHigh"
   TextField "Text field_10" at 7,310 size 53x22; Text 'IW116'
   TextField "Text field_11" at 60,430 size 220x22; Text 'CV-403 - IG Vent Valve Position Fbk'
   IOField "I/O field_16" at 287,430 size 70x22; FormatPattern 999; Unit  %
      ProcessValue <- "12_AI_Data_CV403_SCALED"
   IOField "I/O field_17" at 361,430 size 60x22; FormatPattern 999
   IOField "I/O field_18" at 429,430 size 60x22; FormatPattern 999
   IOField "I/O field_19" at 497,430 size 60x22; FormatPattern 999
   IOField "I/O field_20" at 565,430 size 60x22; FormatPattern 999
   TextField "Text field_12" at 7,430 size 53x22; Text 'IW118'
   TextField "Text field_13" at 60,470 size 220x22; Text 'CA Blower RPM'
   IOField "I/O field_21" at 287,470 size 70x22; FormatPattern 9999; Unit  RPM
      ProcessValue <- "12_AI_Data_E139_RPM_SCALED"
   IOField "I/O field_22" at 361,470 size 60x22; FormatPattern 9999
   IOField "I/O field_23" at 429,470 size 60x22; FormatPattern 9999
   IOField "I/O field_24" at 497,470 size 60x22; FormatPattern 9999
   IOField "I/O field_25" at 565,470 size 60x22; FormatPattern 9999
   TextField "Text field_14" at 7,470 size 54x22; Text 'IW120'
   TextField "Text field_15" at 61,511 size 220x22; Text 'CA Blower Current'
   IOField "I/O field_26" at 288,511 size 70x22; FormatPattern 999.9; Unit  A
      ProcessValue <- "12_AI_Data_E139_AMPS_SCALED"
   IOField "I/O field_27" at 362,511 size 60x22; FormatPattern 9999
   IOField "I/O field_28" at 430,511 size 60x22; FormatPattern 9999
   TextField "Text field_16" at 8,511 size 54x22; Text 'IW122'
   TextField "Text field_17" at 61,552 size 220x22; Text 'LIT-305 - FW Bulk Tank Level'
   IOField "I/O field_31" at 288,552 size 70x22; FormatPattern s99.9; Unit  %
      ProcessValue <- "12_AI_Data_LIT305_SCALED"
   TextField "Text field_18" at 8,552 size 53x22; Text 'IW124'
   TextField "Text field_19" at 61,592 size 220x22; Text 'Spare'
   IOField "I/O field_36" at 288,592 size 70x22; FormatPattern 9.9; Unit  
      ProcessValue <- "12_AI_Data_R1_SPR_AI_126_SCALED"
   IOField "I/O field_37" at 362,592 size 60x22; FormatPattern 9.9
   IOField "I/O field_38" at 430,592 size 60x22; FormatPattern 9.9
   IOField "I/O field_39" at 498,592 size 60x22; FormatPattern 9.9
   IOField "I/O field_40" at 566,592 size 60x22; FormatPattern 9.9
   TextField "Text field_20" at 8,592 size 53x22; Text 'IW126'
   TextField "Text field_21" at 703,151 size 220x22; Text 'Atmospheric Oxygen 1'
   IOField "I/O field_41" at 930,151 size 70x22; FormatPattern 99.99; Unit %
      ProcessValue <- "12_AI_Data_AT_O2_01_SCALED"
   IOField "I/O field_42" at 1004,151 size 60x22; Authorization "Commissioning"; FormatPattern 99.9
      ProcessValue <- "84_Setpoints_AT_O2_1_LowLow"
   IOField "I/O field_43" at 1072,151 size 60x22; Authorization "Commissioning"; FormatPattern 99.9
      ProcessValue <- "84_Setpoints_AT_O2_1_Low"
   IOField "I/O field_44" at 1140,151 size 60x22; FormatPattern 99.9
   IOField "I/O field_45" at 1208,151 size 60x22; FormatPattern 99.9
   TextField "Text field_22" at 650,151 size 53x22; Text 'IW128'
   TextField "Text field_26" at 928,124 size 64x20; Text 'Reading'
   TextField "Text field_27" at 1001,124 size 68x20; Text 'Low Low'
   TextField "Text field_28" at 1082,124 size 37x20; Text 'Low'
   TextField "Text field_29" at 1150,124 size 37x20; Text 'High'
   TextField "Text field_30" at 1203,124 size 74x20; Text 'High High'
   TextField "Text field_31" at 1076,100 size 76x20; Text 'Setpoints'
   TextField "Text field_57" at 703,192 size 220x22; Text 'TIT-315 - Shell CSW Temperature'
   IOField "I/O field_106" at 930,192 size 70x22; FormatPattern s999.9; Unit  °C
      ProcessValue <- "12_AI_Data_TIT315_SCALED"
   IOField "I/O field_107" at 1004,192 size 60x22; FormatPattern s999.9
   IOField "I/O field_108" at 1072,192 size 60x22; FormatPattern s999.9
   TextField "Text field_58" at 650,192 size 54x22; Text 'IW134'
   TextField "Text field_59" at 703,232 size 220x22; Text 'TIT-319 - Inlet CSW Temperature'
   IOField "I/O field_111" at 930,232 size 70x22; FormatPattern s999.9; Unit  °C
      ProcessValue <- "12_AI_Data_TIT319_SCALED"
   IOField "I/O field_112" at 1004,232 size 60x22; FormatPattern s999.9
   IOField "I/O field_113" at 1072,232 size 60x22; FormatPattern s999.9
   TextField "Text field_60" at 650,232 size 53x22; Text 'IW136'
   TextField "Text field_61" at 703,272 size 220x22; Text 'TIT-360 - Outlet CSW Temperature'
   IOField "I/O field_116" at 930,272 size 70x22; FormatPattern s999.9; Unit  °C
      ProcessValue <- "12_AI_Data_TIT360_SCALED"
   IOField "I/O field_117" at 1004,272 size 60x22; FormatPattern s999.9
   IOField "I/O field_118" at 1072,272 size 60x22; FormatPattern s999.9
   TextField "Text field_62" at 650,272 size 53x22; Text 'IW138'
   TextField "Text field_63" at 703,312 size 220x22; Text 'PIT-359 - Inlet CSW Pressure'
   IOField "I/O field_121" at 930,312 size 70x22; FormatPattern 99.9; Unit  Bar
      ProcessValue <- "12_AI_Data_PIT359_SCALED"
   TextField "Text field_64" at 650,312 size 53x22; Text 'IW140'
   TextField "Text field_41" at 133,124 size 89x20; Text 'Description'
   TextField "Text field_42" at 771,124 size 89x20; Text 'Description'
   TextField "Text field_43" at 17,124 size 37x20; Text 'AI'
   TextField "Text field_44" at 661,124 size 37x20; Text 'AI'
   TextField "Text field_47" at 702,352 size 220x22; Text 'PIT-316 - Outlet CSW Pressure'
   IOField "I/O field_81" at 929,352 size 70x22; FormatPattern 99.9; Unit  Bar
      ProcessValue <- "12_AI_Data_PIT316_SCALED"
   TextField "Text field_48" at 649,352 size 53x22; Text 'IW142'
   IOField "I/O field_109" at 1140,192 size 60x22; Authorization "Parameter Change"; FormatPattern s999.9
      ProcessValue <- "84_Setpoints_TIT315_High"
   IOField "I/O field_110" at 1208,192 size 60x22; Authorization "Parameter Change"; FormatPattern s999.9
      ProcessValue <- "84_Setpoints_TIT315_HighHigh"
   IOField "I/O field_114" at 1140,232 size 60x22; Authorization "Parameter Change"; FormatPattern s999.9
      ProcessValue <- "84_Setpoints_TIT319_High"
   IOField "I/O field_115" at 1208,232 size 60x22; Authorization "Parameter Change"; FormatPattern s999.9
      ProcessValue <- "84_Setpoints_TIT319_HighHigh"
   IOField "I/O field_119" at 1140,272 size 60x22; Authorization "Parameter Change"; FormatPattern s999.9
      ProcessValue <- "84_Setpoints_TIT360_High"
   IOField "I/O field_120" at 1208,272 size 60x22; Authorization "Parameter Change"; FormatPattern s999.9
      ProcessValue <- "84_Setpoints_TIT360_HighHigh"
   IOField "I/O field_124" at 1140,312 size 60x22; Authorization "Parameter Change"; FormatPattern 99.9
      ProcessValue <- "84_Setpoints_PIT359_High"
   IOField "I/O field_125" at 1208,312 size 60x22; Authorization "Parameter Change"; FormatPattern 99.9
      ProcessValue <- "84_Setpoints_PIT359_HighHigh"
   IOField "I/O field_84" at 1139,352 size 60x22; Authorization "Parameter Change"; FormatPattern 99.9
      ProcessValue <- "84_Setpoints_PIT316_High"
   IOField "I/O field_85" at 1207,352 size 60x22; Authorization "Parameter Change"; FormatPattern 99.9
      ProcessValue <- "84_Setpoints_PIT316_HighHigh"
   IOField "I/O field_122" at 1004,312 size 60x22; Authorization "Parameter Change"; FormatPattern 99.9
      ProcessValue <- "84_Setpoints_PIT359_LowLow"
   IOField "I/O field_123" at 1072,312 size 60x22; Authorization "Parameter Change"; FormatPattern 99.9
      ProcessValue <- "84_Setpoints_PIT359_Low"
   IOField "I/O field_82" at 1003,352 size 60x22; Authorization "Parameter Change"; FormatPattern 99.9
      ProcessValue <- "84_Setpoints_PIT316_LowLow"
   IOField "I/O field_83" at 1071,352 size 60x22; Authorization "Parameter Change"; FormatPattern 99.9
      ProcessValue <- "84_Setpoints_PIT316_Low"
   TextField "Text field_52" at 17,91 size 333x26; Text 'IGG Control System PLC (Rack 1)'
   TextField "Text field_54" at 649,719 size 228x62; Text 'Note: CSW = Cooling Sea Water'
   Button "Button_1" at 1160,732 size 100x35; TextOn 'BWTS Digital Inputs.'; TextOff 'Next'
      on Click: ActivateScreen("BC Analogue Inputs", 0)
   TextField "Text field_25" at 60,231 size 220x22; Text 'PIT-102 - CA Pressure (Post-Ignition)'
   IOField "I/O field_52" at 361,231 size 60x22; Authorization "Parameter Change"; FormatPattern 9999
      ProcessValue <- "84_Setpoints_PIT102_Post_LowLow"
   IOField "I/O field_53" at 429,231 size 60x22; Authorization "Parameter Change"; FormatPattern 9999
      ProcessValue <- "84_Setpoints_PIT102_Post_Low"
   IOField "I/O field_54" at 497,231 size 60x22; Authorization "Parameter Change"; FormatPattern 9999
      ProcessValue <- "84_Setpoints_PIT102_Post_High"
   IOField "I/O field_55" at 565,231 size 60x22; Authorization "Parameter Change"; FormatPattern 9999
      ProcessValue <- "84_Setpoints_PIT102_Post_HighHigh"
   TextField "Text field_32" at 7,231 size 53x22; Text 'IW112'
   TextField "Text field_33" at 60,391 size 220x22; Text 'PIT-402 - IG Outlet Pres. (Post-Ignitn)'
   IOField "I/O field_57" at 361,391 size 60x22; Authorization "Parameter Change"; FormatPattern 9999
      ProcessValue <- "84_Setpoints_PIT402_Post_LowLow"
   IOField "I/O field_58" at 429,391 size 60x22; Authorization "Parameter Change"; FormatPattern 9999
      ProcessValue <- "84_Setpoints_PIT402_Post_Low"
   IOField "I/O field_59" at 497,391 size 60x22; Authorization "Parameter Change"; FormatPattern 9999
      ProcessValue <- "84_Setpoints_PIT402_Post_High"
   IOField "I/O field_60" at 565,391 size 60x22; Authorization "Parameter Change"; FormatPattern 9999
      ProcessValue <- "84_Setpoints_PIT402_Post_HighHigh"
   TextField "Text field_34" at 7,391 size 53x22; Text 'IW116'
   TextField "Text field_35" at 61,191 size 220x22; Text 'PIT-102 - CA Pressure (Main)'
   IOField "I/O field_50" at 362,191 size 60x22; Authorization "Parameter Change"; FormatPattern 9999
      ProcessValue <- "84_Setpoints_PIT102_Main_LowLow"
   IOField "I/O field_63" at 430,191 size 60x22; Authorization "Parameter Change"; FormatPattern 9999
      ProcessValue <- "84_Setpoints_PIT102_Main_Low"
   IOField "I/O field_64" at 498,191 size 60x22; Authorization "Parameter Change"; FormatPattern 9999
      ProcessValue <- "84_Setpoints_PIT102_Main_High"
   IOField "I/O field_65" at 566,191 size 60x22; Authorization "Parameter Change"; FormatPattern 9999
      ProcessValue <- "84_Setpoints_PIT102_Main_HighHigh"
   TextField "Text field_36" at 8,191 size 53x22; Text 'IW112'
   TextField "Text field_37" at 61,349 size 220x22; Text 'PIT-402 - IG Outlet Pres. (Main)'
   IOField "I/O field_69" at 362,349 size 60x22; Authorization "Parameter Change"; FormatPattern 9999
      ProcessValue <- "84_Setpoints_PIT402_Main_LowLow"
   IOField "I/O field_70" at 430,349 size 60x22; Authorization "Parameter Change"; FormatPattern 9999
      ProcessValue <- "84_Setpoints_PIT402_Main_Low"
   IOField "I/O field_71" at 498,349 size 60x22; Authorization "Parameter Change"; FormatPattern 9999
      ProcessValue <- "84_Setpoints_PIT402_Main_High"
   IOField "I/O field_72" at 566,349 size 60x22; Authorization "Parameter Change"; FormatPattern 9999
      ProcessValue <- "84_Setpoints_PIT402_Main_HighHigh"
   TextField "Text field_38" at 8,349 size 53x22; Text 'IW116'
   IOField "I/O field_29" at 566,511 size 60x22; FormatPattern 9999
   IOField "I/O field_30" at 499,511 size 60x22; FormatPattern 9999
   IOField "I/O field_32" at 361,552 size 60x22; FormatPattern 9999
   IOField "I/O field_33" at 429,552 size 60x22; FormatPattern 9999
   IOField "I/O field_34" at 565,552 size 60x22; FormatPattern 9999
   IOField "I/O field_35" at 498,552 size 60x22; FormatPattern 9999
   TextField "Text field_39" at 1109,687 size 151x62; Text 'To BC Analogue Inputs'
   AlarmView "Alarm view_1" at 0,777 size 1280x23
   Group "Group" at 455,41 size 373x50
   Button "HmiScreenItemData_8" at 469,45 size 355x40; TextOn 'Back'; TextOff 'Text'
   TextField "Screen title" at 455,41 size 373x50; Text 'Screen title'